   REGION R-trig
       #RTIRG_iReset(CLK := #iReset);
       #RTRIG_iFailSafe(CLK := #iFailSafe);
       #RTIRG_jog(CLK := #iJogOpen XOR #iJogClose);
       #RTIRG_auto(CLK := NOT #iMan);
       #RTRIG_iFailSafe_released(CLK := #iFailSafe);
       #RTRIG_iInterlook_released(CLK := #iInterlook);
       #RTRIG_jogOpen_released(CLK := NOT #iJogOpen);
       #RTRIG_jogClose_released(CLK := NOT #iJogClose);
   END_REGION

   REGION Timeout  

       // Quick timeout:
       // Cheak at intervals that the position moves towards the setpoint.
       // This give a quicker feedback, then the long timeout.
       IF #action <> #old.action
           OR #RTIRG_jog.Q
           OR #RTRIG_iFailSafe.Q
       THEN
           RESET_TIMER(#TONR_quckTimeoutInterval);
           #quickTimeoutLastPos := #io.in.pos;
       ELSIF #action <> #NO_ACTION AND #conf.quickTimeoutEnable THEN
           // Quick timeout in action.
           #TONR_quckTimeoutInterval.TONR(IN := #io.out.open OR #io.out.close,
                                          PT := #conf.quickTimeoutIntervalCheaks);
           IF #TONR_quckTimeoutInterval.Q THEN
               // A new interval check, now see if the valve has moved sufficient.
               #out.qucikTimeout :=
               ABS(#quickTimeoutLastPos - #io.in.pos) < #conf.qucikTimeoutMinMovement;
               RESET_TIMER(#TONR_quckTimeoutInterval);
               // Only store the old value if the valve has done progress towards the SP.
               IF #action = #OPEN AND #io.in.pos > #quickTimeoutLastPos
                   OR #action = #CLOSE AND #io.in.pos < #quickTimeoutLastPos
               THEN
                   #quickTimeoutLastPos := #io.in.pos;
               END_IF;
           END_IF;
       END_IF;

       // Long timeout:
       // Max time the valve can operate before timeout, and the valve will stop.
       #TONR_timeout.TONR(IN := #io.out.open OR #io.out.close,
                          PT := #conf.longTimeout,
                          Q => #out.longTimeout);
       // Reset timeout
       IF #RTIRG_iReset.Q
           OR #RTRIG_iFailSafe.Q
           OR #conf.autoReset AND (
           (* *)#RTIRG_jog.Q
           (* *)OR #iSP <> #old.SP AND #iMan
           (* *)OR #RTIRG_jog.Q)
       THEN
           RESET_TIMER(#TONR_timeout);
           RESET_TIMER(#TONR_quckTimeoutInterval);
           #out.qucikTimeout := false;
           #qTimeout := false;
       END_IF;
   END_REGION

   REGION Decide
       // Decide what to do ...

       // Error, timeout, failSafe and Interlook.
       IF #TONR_timeout.Q THEN
           #action := #NO_ACTION;
       ELSIF #iFailSafe THEN
           // Timeout will be reseted once if iFailSafe is activated.
           #action := #conf.feilSafeAction;
       ELSIF #iStop
           // If pos.error and there are not end-limit-switces.
           OR #io.in.posError AND (#conf.simFullyOpenWithPos OR #conf.simFullyClosedWithPos)
           OR #out.qucikTimeout
           OR #RTRIG_jogOpen_released.Q
           OR #RTRIG_jogClose_released.Q
           OR #iExternalError
       THEN
           #action := #NO_ACTION;

           // ==========================================================================
           // JOG-mode
       ELSIF #iJogOpen XOR #iJogClose THEN
           // Open or close the valve little by little. When either of the jog
           // inputs are true. This way of controlling the valve has priority
           // over setpoint (bellow).
           RESET_TIMER(#TON_regModeWait);
           IF #iJogOpen THEN
               #action := #OPEN;
           ELSIF #iJogClose THEN
               #action := #CLOSE;
           END_IF;
       ELSIF #io.in.posError THEN
           #action := #NO_ACTION;
       ELSE
           // ==========================================================================
           // SP-mode:
           // Controll the valve by a setpoint, using the feedback position to 
           // determined if the valve should open or close. SP should be given in percent.

           IF (#iSP <> #old.SP // SP has changed.
               OR #RTIRG_auto.Q // Auto has just been enabled, and the valve is out of pos.
               (* *)AND ABS(#iSP - #io.in.pos) > #conf.regModeMinOffset
               OR NOT #iMan AND ( // In auto
               (* *)#RTIRG_iReset.Q // Avoid dead lock
               (* *)OR #RTRIG_iFailSafe_released.Q
               (* *)OR #RTRIG_iInterlook_released.Q
               (* *)OR #RTRIG_jogClose_released.Q OR #RTRIG_jogOpen_released.Q )
               (* *)) AND (
               (*     *)NOT #iRegMode // Not regMode, no aditional requirements.
               (*     *)OR #TON_regModeWait.Q AND ( // A break between each move.
               (*        *)// Offset is bigger then a certain offset.
               (*        *)ABS(#iSP - #io.in.pos) > #conf.regModeMinOffset
               (*        *)// At almost closed and open, the offset requirement
               (*        *)// may not be fulfilled.
               (*        *)OR #io.in.pos > #conf.fullyOpenPosLim - #conf.endPosWithoutPreStop
               (*        *)OR #io.in.pos < #conf.endPosWithoutPreStop))
               // regMode should be used when a valve is controlled by a PID.
               // When the valve is in regMode, then there will be a time break between each 
               // movment. And there is a need a certain offset before an ajustment is done.
               // This behavior significantly prevents wear on the valve. If the valve is not
               // in regMode, then each change in SP will make the valve operate.
           THEN
               IF #iSP > #io.in.pos THEN
                   #action := #OPEN;
               ELSIF #iSP < #io.in.pos THEN
                   #action := #CLOSE;
               END_IF;
           END_IF;

           // --------------------------------------
           // SP-reached-pos:
           // 
           // In the main area where the valve operate, it will shut off the outputs, a
           // tiny bit before it reach the SP. This make the valve, stop exacly on SP.
           // In the area of almost closed and almost open this function is disable,
           // this makes sure that it's possible to open or close the valve entirly.
           #pre := SEL(G := #iSP > #conf.fullyOpenPosLim - #conf.endPosWithoutPreStop
                       OR #iSP < #conf.endPosWithoutPreStop,
                       IN0 := #conf.preStop, IN1 := 0);
           // Detect reached position
           IF #action = #OPEN AND (#io.in.pos > #iSP - #pre OR #io.in.fullyOpen)
               OR #action = #CLOSE AND (#io.in.pos < #iSP + #pre OR #io.in.fullyClosed)
           THEN
               #action := #NO_ACTION;
               RESET_TIMER(#TON_regModeWait);
           END_IF;
       END_IF;
       // In regMode this timer need to finnish before a new movement can be done.
       #TON_regModeWait.TON(IN := true,
                            PT := #conf.regModeTimeBreak);
   END_REGION

   REGION Gentle
       // If a big valve closes or open to fast, it can damage the pipes or other
       // equipment. This section make time breaks on closing or opening. 

       #gentleMode := #io.in.pos < #conf.gentleActivteLowLimit // ->
       // -> The function is only active under a ceratain position limit.
       AND (NOT #iFailSafe OR #conf.gentleAlsoOnFailSafe)
       // AlsoOnFailSafe: It's possible to disable the function for emergencies
       // by setting the value false.
       AND (#conf.gentleOpenEnable AND #action = #OPEN
       (* *)OR #conf.gentleCloseEnable AND #action = #CLOSE);    

       // The time break will increase as the valve move from the limit towards close.
       #pause := REAL_TO_DINT(#conf.gentleTimePauseBias
                              + (#io.in.pos / #conf.gentleActivteLowLimit)
                              * #conf.gentleTimePauseDelta);
       IF #gentleMode THEN
           #TON_gentle.TON(IN := true,
                           PT := SEL(G := #gentleAction, // Toggle times
                                     IN0 := #conf.gentleTimeRun,
                                     IN1 := #pause));
           IF #TON_gentle.Q THEN
               #gentleAction := NOT #gentleAction;
               RESET_TIMER(#TON_gentle); 
           END_IF;
           #action2 := SEL(G := #gentleAction, // Toggle action
                           IN0 := #action, IN1 := #NO_ACTION);
       ELSE
           RESET_TIMER(#TON_gentle);
           #gentleAction := false;
           // If the carefully-function is disabled, then just forward
           // the action value to the next stage.
           #action2 := #action;
       END_IF;
   END_REGION

   REGION Output
       // Make a smal time break when valve change direction. This make sure that
       // that both outputs are not active at the same time.
       #TP_toggleOut.TP(IN := #action2 <> #old.action2 AND #old.action2 <> #NO_ACTION,
                        PT := #conf.toggleTimeBreak);

       // Outputs
       IF #TP_toggleOut.Q THEN // A small time break.
           #io.out.open := false;
           #io.out.close := false;
       ELSIF #iFailSafe 
           OR #iJogClose OR #iJogOpen
       THEN
           // When failSafe or jog is active both the limit-switch and positon
           // signal most indicate that the valve is in correct position. This
           // in case one of the signals isn't working.
           #io.out.open := #action2 = #OPEN AND NOT #bothSensors.open;
           #io.out.close := #action2 = #CLOSE AND NOT #bothSensors.closed;
       ELSIF #iInterlook THEN
           #io.out.open := false;
           #io.out.close := false;
       ELSE
           #io.out.open := #action2 = #OPEN AND NOT #io.in.fullyOpen;
           #io.out.close := #action2 = #CLOSE AND NOT #io.in.fullyClosed;
       END_IF;
   END_REGION

   REGION Old    
       // Store values, to check if they has changed until next scan.
       #old.SP := #iSP;
       #old.action := #action;
       #old.action2 := #action2;
   END_REGION

   #qTimeout := #out.qucikTimeout OR #out.longTimeout;
END_FUNCTION_BLOCK

FUNCTION_BLOCK "motorValve"   // FB10, SCL
{ S7_Optimized_Access := 'TRUE' }
VERSION : 0.1
   VAR_INPUT
      iFeedbackPosition : Real;
      iFeddbackPosError : Bool;
      iFeedbackFullyOpen : Bool;
      iFeedbackFullyClosed : Bool;
   END_VAR
   VAR_OUTPUT
      qOpen : Bool;
      qClose : Bool := FALSE;
   END_VAR
   VAR RETAIN
      hmi : "motorValveHmiUdt";
   END_VAR
   VAR
      valve : "motorValveCtrl";
      SP : Real;
      SP_auto : Real;
   END_VAR
   VAR CONSTANT
      AUTO : SInt := 0;
      MAN_LOCAL : SInt := 1;
      MAN_REMOTE : SInt := 2;
   END_VAR
BEGIN
   // Valve with analog feedback.

   REGION Simulation
       IF #hmi.sim.enable AND NOT #valve.iFailSafe THEN
           // Simulation of input signal, not possible if in fail safe mode.
           #hmi.io.in.pos := #hmi.sim.pos;
           #hmi.io.in.posError := false;
           #hmi.io.in.fullyOpen := #hmi.sim.pos > #hmi.conf.fullyOpenPosLim;
           #hmi.io.in.fullyClosed := #hmi.sim.pos < #hmi.conf.fullyClosedPosLim;
       ELSE
           // Input mapping
           #hmi.io.in.pos := #iFeedbackPosition;
           #hmi.io.in.posError := #iFeddbackPosError;
           #hmi.io.in.fullyOpen := #iFeedbackFullyOpen;
           #hmi.io.in.fullyClosed := #iFeedbackFullyClosed;
       END_IF;
   END_REGION

   REGION Man / auto    
       IF #hmi.cmd.stop THEN
           #hmi.autoMan := #MAN_LOCAL;
       ELSIF #hmi.cmd.jogOpen XOR #hmi.cmd.jogClose THEN
           #hmi.autoMan := #MAN_LOCAL;
           #SP := #iFeedbackPosition;
       ELSIF #hmi.cmd.openFully XOR #hmi.cmd.closeFully THEN
           #hmi.autoMan := #MAN_LOCAL;
           #SP := SEL(G := #hmi.cmd.openFully, IN0 := 0, IN1 := 100);
       ELSIF #hmi.autoMan = #MAN_LOCAL THEN
           #SP := #hmi.SP;
       ELSIF #hmi.autoMan = #AUTO THEN
           #SP := #SP_auto;
           // If auto is controlled by a pid then #hmi.conf.regMode need to be enabled.
       END_IF;
       #hmi.SP := #valve.iSP := #SP_auto := #SP;
       // Forward auto or man to the valve controller.
       CASE #hmi.autoMan OF
           #MAN_LOCAL, #MAN_REMOTE:
               #valve.iMan := true;
           #AUTO:
               #valve.iMan := false;
       END_CASE;
   END_REGION

   REGION Valve controller.        
       // Main valve controller block.
       #valve(// iFailSafe
              // iInterlook
              // iRegMode
              iStop := #hmi.cmd.stop,
              iJogOpen := #hmi.cmd.jogOpen,
              iJogClose := #hmi.cmd.jogClose,
              iReset := #hmi.cmd.reset,
              qTimeout => #hmi.error.timeout,
              conf := #hmi.conf,
              io := #hmi.io);
       #qOpen := #hmi.io.out.open; // Outputs
       #qClose := #hmi.io.out.close;
   END_REGION

   REGION Position error    
       #hmi.error.posError :=
       #iFeedbackFullyOpen AND #iFeedbackFullyClosed
       OR #iFeedbackFullyOpen
       (* *)AND #iFeedbackPosition < #hmi.conf.fullyOpenPosLim - #hmi.conf.regModeMinOffset
       (* *)AND NOT #hmi.conf.simFullyOpenWithPos
       OR #iFeedbackFullyClosed
       (* *)AND #iFeedbackPosition > #hmi.conf.fullyClosedPosLim + #hmi.conf.regModeMinOffset
       (* *)AND NOT #hmi.conf.simFullyClosedWithPos;
   END_REGION

   REGION End
       // Count secounds the valve has been operating, and number of starts.
       "operatingTime"(in := #qOpen OR #qClose,
                       opr := #hmi.operatingTime);

       // Reset signals.
       #hmi.cmd.jogOpen := false;
       #hmi.cmd.jogClose := false;
       #hmi.cmd.openFully := false;
       #hmi.cmd.closeFully := false;
       #hmi.cmd.reset := false;
       #hmi.cmd.man := false;
       #hmi.cmd.auto := false;
       CASE #hmi.autoMan OF // Reset stop signal, only if in man.
           #MAN_LOCAL, #MAN_REMOTE: // If in auto, then do nothing.
               #hmi.cmd.stop := false;
       END_CASE;

       // Other signals to HMI
       #hmi.info.failSafe := #valve.iFailSafe;
       #hmi.info.interlook := #valve.iInterlook;
       #hmi.info.regMode := #valve.iRegMode;

       #hmi.sim.simByPlc := #hmi.io.simulated;
       #hmi.io.simulated := false;
   END_REGION
END_FUNCTION_BLOCK

FUNCTION_BLOCK "motorValveSimulation"   // FB20, SCL
{ S7_Optimized_Access := 'TRUE' }
VERSION : 0.1
   VAR_INPUT
      speed : Real := 1.0;
   END_VAR
   VAR_IN_OUT
      io : "motorValveIoUdt";
   END_VAR
   VAR
      old : UDInt;
      sn : UDInt;
   END_VAR
   VAR_TEMP
      t : DTL;
      "e" : Int;
   END_VAR
BEGIN
   #"e" := RD_SYS_T(#t);
   #sn := #t.NANOSECOND / 100000 + #t.SECOND * 10;

   IF #sn = #old THEN
       IF #io.out.open THEN
           #io.in.pos += #speed * 0.1;
       ELSIF #io.out.close THEN
           #io.in.pos -= #speed;
       END_IF;
   END_IF;
   #old := #sn;

   #io.in.pos := LIMIT(MN := 0, IN := #io.in.pos, MX := 100);
   #io.in.fullyOpen := #io.in.pos > 99;
   #io.in.fullyClosed := #io.in.pos < 1;

   #io.simulated := true;
END_FUNCTION_BLOCK

FUNCTION "ioGlobalMotorValveLinking" : Void   // FC24, SCL
{ S7_Optimized_Access := 'TRUE' }
VERSION : 0.1
   VAR_IN_OUT
      ioGlobal : "ioGlobal_FB";
      valve : "motorValve";
   END_VAR
BEGIN
   // Link ioGlobal with valve functions.

   // A id for each io
   #ioGlobal.z.ioIdCnt += 1;

   IF #ioGlobal.info2ioBlocks.disableAllSim THEN
       #valve.hmi.sim.enable := false;
   END_IF;
   // Count active simulations
   #ioGlobal.collectInfo.activeSimCnt +=
   BOOL_TO_UINT(#valve.hmi.sim.enable OR #valve.hmi.sim.simByPlc);

   // Count number of errors
   #ioGlobal.collectInfo.errorCnt +=
   BOOL_TO_UINT(#valve.hmi.io.in.posError OR #valve.hmi.error.timeout);
END_FUNCTION

// folder: Library/Valves/Blocks and UDT's/z Dev

FUNCTION_BLOCK "motorValveDigital"   // FB11, SCL
{ S7_Optimized_Access := 'TRUE' }
VERSION : 0.1
   VAR_INPUT
      iAction : SInt;   // 0=no-action, 1=Open, 2=Close
      iFailSafe : Bool;   // Open or close the valve entirly, set inside conf.
      iInterlook : Bool;   // Stop movement, valve will continue when input is set back false.
      iStop : Bool;   // Stop movement, also after var. is back false.
      iJogOpen : Bool;   // Move the valve towards open when true, has priority over SP.
      iJogClose : Bool;   // Move the valve towards close when true, has priority over SP.
      iReset : Bool;   // Reset timeout.
   END_VAR
   VAR_OUTPUT
      qTimeout : Bool;   // (quick and long timeout)
   END_VAR
   VAR
      action : SInt;   // 1=open, 2=close
      actionOut : SInt;
      oldAction : SInt;
      oldActionOut : SInt;
      RTIRG_iFailSafe : R_TRIG;
      RTIRG_iReset : R_TRIG;
      RTIRG_jog : R_TRIG;
      TP_toggleOut : IEC_TIMER;
      TON_gentle : IEC_TIMER;
      TONR_gentle : IEC_TIMER;
      TONR_timeout : IEC_TIMER;
      TON_regModeWait : IEC_TIMER;
      gentleAction : Bool;
   END_VAR
   VAR_TEMP
      reset : Bool;
   END_VAR
   VAR CONSTANT
      NO_ACTION : SInt := 0;
      OPEN : SInt := 1;
      CLOSE : SInt := 2;
   END_VAR
BEGIN
   // #conf - "motorValveConfUdt"
   // #io - "motorValveIoUdt"

   // Valve 

   (*

   //R-TRIG'S
   #RTIRG_iReset(CLK := #iReset);
   #RTIRG_iFailSafe(CLK := #iFailSafe); // Reset timeout once on failSafe.
   #RTIRG_jog(CLK := #iJogOpen XOR #iJogClose);

   REGION Timeout-and-reset
       // Max time the valve can operate before timeout, and the valve will stop.
       #TONR_timeout.TONR(IN := #io.out.open OR #io.out.close,
                          PT := #conf.longTimeout,
                          Q => #qTimeout);

       // Reset timeout
       IF #iJogOpen OR #iJogClose THEN
           #reset := #RTIRG_jog.Q AND (#conf.autoReset OR NOT #qTimeout);
       END_IF;
       IF #RTIRG_iReset.Q OR #RTIRG_iFailSafe.Q OR #reset THEN
           RESET_TIMER(#TONR_timeout);
           #qTimeout := false;
       END_IF;
   END_REGION

   REGION Decide
       // Error, timeout, failSafe and Interlook.
       IF #TONR_timeout.Q THEN
           #action := #NO_ACTION;
       ELSIF #iFailSafe THEN // Timeout will be reseted once if iFailSafe is activated.
           #action := #conf.feilSafeAction;
       ELSIF #iStop THEN
           #action := #NO_ACTION;
           // ==========================================================================
           // JOG-mode
       ELSIF #iJogOpen OR #iJogClose THEN
           // Open or close the valve little by little. When either of the jog
           // inputs are true. This way of controlling the valve has priority
           // over setpoint (bellow).
           RESET_TIMER(#TON_regModeWait);
           IF #iJogOpen AND #iJogClose THEN
               #action := #NO_ACTION;
           ELSIF #iJogOpen THEN
               #action := #OPEN;
           ELSIF #iJogClose THEN
               #action := #CLOSE;
           ELSE
               ;
           END_IF;
       END_IF;
   END_REGION

   REGION Gentle
       // If a big valve closes or open to fast, it can damage the pipes or other
       // equipment. This section make time breaks on closing or opening. 
       IF #io.in.pos < #conf.gentleActivteLowLimit // ->
           // -> The function is only active under a ceratain position limit.
           AND (NOT #iFailSafe OR #conf.gentleAlsoOnFailSafe)
           // AlsoOnFailSafe: It's possible to disable the function for emergencies
           // by setting the value false.
           AND (#conf.gentleOpenEnable AND #action = #OPEN
           (* *)OR #conf.gentleOpenEnable AND #action = #CLOSE)
       THEN
           #TON_gentle.PT := SEL(G := #gentleAction, // Toggle times
                                 IN0 := #conf.gentleTimeRun,
                                 IN1 := #conf.gentleTimePauseBias);
           #TON_gentle.TON(IN := true,
                           PT := #TON_gentle.PT);
           IF #TON_gentle.Q THEN
               #gentleAction := NOT #gentleAction;
               RESET_TIMER(#TON_gentle);
           END_IF;
           #actionOut := SEL(G := #gentleAction, // Toggle action
                             IN0 := #action, IN1 := #NO_ACTION);
       ELSE
           RESET_TIMER(#TON_gentle);
           #gentleAction := false;
           // If the carefully-function is disabled, then just forward
           // the action value to the next stage.
           #actionOut := #action;
       END_IF;
   END_REGION

   REGION Output
       // Make a smal time break when valve change direction. This make sure that
       // that both outputs are not active at the same time.
       #TP_toggleOut.TP(IN := #actionOut <> #oldActionOut AND #oldActionOut <> #NO_ACTION,
                        PT := #conf.toggleTimeBreak);
       // Outputs
       IF #TP_toggleOut.Q THEN
           #io.out.open := false;
           #io.out.close := false;
       ELSIF #iFailSafe THEN
           #io.out.open := #conf.feilSafeAction = #OPEN AND NOT #io.in.fullyOpen;
           #io.out.close := #conf.feilSafeAction = #CLOSE AND NOT #io.in.fullyClosed;
       ELSIF #iInterlook OR #iStop THEN
           #io.out.open := false;
           #io.out.close := false;
       ELSE
           #io.out.open := #actionOut = #OPEN AND NOT #io.in.fullyOpen;
           #io.out.close := #actionOut = #CLOSE AND NOT #io.in.fullyClosed;
       END_IF;
   END_REGION

   REGION Old
       #oldAction := #action;
       #oldActionOut := #actionOut;
   END_REGION


   // *)
END_FUNCTION_BLOCK

FUNCTION_BLOCK "motorValveAproxPos"   // FB24, SCL
{ S7_Optimized_Access := 'TRUE' }
VERSION : 0.1
   VAR_IN_OUT
      io : "motorValveIoUdt";
   END_VAR
   VAR
      conf : Struct
         maxAvoid : Real := 4.0;
      END_STRUCT;
      oldSecAndMsec10 : UInt;
      posPrT : UInt;
      "timer" : IEC_TIMER;
      first_scan : Bool := TRUE;
      RTRIG_fullyOpen : R_TRIG;
      RTRIG_fullyClosed : R_TRIG;
      rangeTime : Time;
      tries : Array[0..7] of Time;
   END_VAR
   VAR_TEMP
      "e" : Int;
      rd_sys_t : DTL;
      secAndMsec10 : UInt;
      sPos : Int;
      t : Int;
      c : Int;
      mx : Time;
      mn : Time;
   END_VAR
BEGIN
   // #io - "motorValveIoUdt"


   // For valve without position sensor. Calculate the position based on long
   // time the valve has been opening and closing.

   (* FUNCTION NOT FINISHED...

   #e := RD_SYS_T(#rd_sys_t);
   #secAndMsec10 := #rd_sys_t.SECOND * 100 + UDINT_TO_UINT(#rd_sys_t.NANOSECOND / 10000);
   #t := USINT_TO_INT( (#secAndMsec10 - #oldSecAndMsec10 + 6000) MOD 6000);
   #oldSecAndMsec10 := #secAndMsec10;

   #io.in.posError := #io.in.posError AND NOT #first_scan;

   #RTRIG_fullyOpen(CLK := #io.in.fullyOpen);
   #RTRIG_fullyClosed(CLK := #io.in.fullyClosed);

   IF #RTRIG_fullyOpen.Q OR #RTRIG_fullyClosed.Q THEN
       RESET_TIMER(#timer);
       #timer.PT := T#10m;
   END_IF;



   #c := 7 - 1;
   WHILE #c >= 0 DO
       #tries[#c + 1] := #tries[#c];
       #c -= 1;
   END_WHILE;
   #tries[0] := T#123s;

   #mn := T#24d;
   FOR #c := 1 TO 6 BY 2 DO
       #mx := MAX(IN1 := #tries[#c], IN2 := #mx);
       #mn := MIN(IN1 := #tries[#c], IN2 := #mn);
   END_FOR;
   // #mx - #mn ;

   (*IF #first_scan THEN
       #io.in.posError := true;
   END_IF;*)


   IF #io.out.open XOR #io.out.close THEN
       #sPos := SEL(G := #io.out.close, IN0 := #sPos + #t, IN1 := #sPos - #t);
   END_IF;


   // #io.in.pos

   #first_scan := false;

   *)
END_FUNCTION_BLOCK

// folder: Library/Valves/Puls valve

FUNCTION_BLOCK "pulsValve"   // FB25, SCL
{ S7_Optimized_Access := 'TRUE' }
VERSION : 0.1
   VAR_INPUT
      iOpening : Bool;
      iCloses : Bool;
      iPuls : Bool;
      iFullyOpen : Bool;
      iFullyClosed : Bool;
      iConfTimeout : Time := T#3S;
      iConfPulsesBetweenOpenAndClosed : Int;
   END_VAR
   VAR_OUTPUT
      qPos : Real;
      qUnknownPos : Bool;
   END_VAR
   VAR
      cnt : Int;
      rtrig_puls : R_TRIG;
      "timer" : IEC_TIMER;
      first_scan : Bool := TRUE;
   END_VAR
   VAR CONSTANT
      NUMBER_PULES_NOT_CONFIGERED : Int := 0;
   END_VAR
BEGIN
   // Valve position based on puls feedback 

   #rtrig_puls(CLK := #iPuls);
   #"timer".TON(IN := (#iOpening OR #iCloses) AND NOT #rtrig_puls.Q,
              PT := #iConfTimeout);
   IF #iConfPulsesBetweenOpenAndClosed = 0 // Number of pules not configured
       OR #"timer".Q
       OR #first_scan  // 
   THEN
       #qUnknownPos := true;
   ELSIF #iFullyOpen THEN
       #cnt := #iConfPulsesBetweenOpenAndClosed;
       #qUnknownPos := false;
   ELSIF #iFullyClosed THEN
       #cnt := 0;
       #qUnknownPos := false;
   ELSE
       IF #iOpening AND #iCloses THEN
           ; // No action
       ELSIF #rtrig_puls.Q THEN
           #cnt += BOOL_TO_INT(#iOpening);
           #cnt -= BOOL_TO_INT(#iCloses);
       END_IF;
   END_IF;
   #qPos := INT_TO_REAL(#cnt) / INT_TO_REAL(#iConfPulsesBetweenOpenAndClosed) * 100;
   #first_scan := false;
END_FUNCTION_BLOCK

// folder: Library/sys/Generate User Msg

FUNCTION_BLOCK "genUsrMsg"   // FB3, SCL
{ S7_Optimized_Access := 'TRUE' }
VERSION : 0.1
   VAR_INPUT
      TextID : UInt;
   END_VAR
   VAR
      TextListID : UInt;
      outgoingAlarm : Bool;   // false: Incoming alarm.
      assocValues : Array[3..10] of UInt;
      "e" : Int;
   END_VAR
   VAR_TEMP
      tmpAssocValues : AssocValues;
      c : Int;
   END_VAR
BEGIN
   // Generate user diagnostic alarms 

   // #assocValues 1 and 2 allready in use by instruction.
   FOR #c := 3 TO 10 DO
       #tmpAssocValues.Value[#c] := #assocValues[#c];
   END_FOR;

   #"e" := Gen_UsrMsg
   (Mode := 1 + BOOL_TO_UINT(#outgoingAlarm)
    ,// 1: incoming alarm. 2: outgoing alarm.
    TextID := #TextID,
   TextListID := #TextListID, // (Right click and show collom-id) 
    AssocValues := #tmpAssocValues);

   (* Assoc Values:

   "This is a usr. msg: @3I%6d@"  // Assoc val 3, 6 digits. (1st val)
   "This is an other usr. msg: @5I%6d@"  // Assoc val 5, 6 digits.

   *)
END_FUNCTION_BLOCK

FUNCTION_BLOCK "example_genUsrMsg"   // FB8, SCL
{ S7_Optimized_Access := 'TRUE' }
VERSION : 0.1
   VAR
      Gen_UsrMsg : "genUsrMsg";
      some_error : Bool;
   END_VAR
BEGIN
   #Gen_UsrMsg.TextListID := 512; // See PLC alarm text lists.

   IF #some_error THEN
       #Gen_UsrMsg(1); // Text id for this alarm 
   END_IF;
END_FUNCTION_BLOCK

// ===== library types =====

TYPE "timeFormatUdt"
   STRUCT
      OFF : SInt := 0;
      MILLISECOND : SInt := 1;
      SECOUNDS : SInt := 2;
      MINUTES : SInt := 3;
      HOURS : SInt := 4;
      DAYS : SInt := 5;
   END_STRUCT;
END_TYPE

// folder: Library/Conversion/time_to_str

FUNCTION "str::" : String   // FC30, SCL
{ S7_Optimized_Access := 'TRUE' }
VERSION : 0.1
   VAR_INPUT
      in : Time;   // Time to be converted in to string.
   END_VAR
   VAR_TEMP
      t : DTL;
      dayOrHour : Bool;
   END_VAR
BEGIN
   // Time to string.

   #t += #in; // Implicit convert to dtl.
   #t.DAY -= 1; 
   #tStr := ''; 

   IF #t.DAY <> 0 THEN
       #tStr := CONCAT(IN1 := RIGHT
                              (IN := S_CONV(#t.DAY),
                               L := 1 + BOOL_TO_INT(#t.DAY > 9)),
                              IN2 := ', ');
   END_IF;
   IF #t.HOUR <> 0 OR LEN(#tStr) <> 0 THEN
       #tStr := CONCAT(IN1 := #tStr,
                              IN2 := RIGHT
                              (IN := S_CONV(#t.HOUR),
                               L := 1 + BOOL_TO_INT(#t.HOUR > 9)),
                              IN3 := ':');
   END_IF;
   #tStr := CONCAT(IN1 := #tStr,
                          IN2 := RIGHT
                          (IN := S_CONV(#t.MINUTE),
                           L := 1 + BOOL_TO_INT(#t.MINUTE > 9)),
                          IN3 := ':');
   #tStr := CONCAT(IN1 := #tStr,
                          IN2 := RIGHT
                          (IN := S_CONV(#t.SECOND),
                           L := 1 + BOOL_TO_INT(#t.SECOND > 9)));

   // https://github.com/rexhip/
END_FUNCTION

// folder: Library/State machine

FUNCTION "sTimer" : Bool   // FC23, SCL
{ S7_Optimized_Access := 'TRUE' }
VERSION : 0.1
   VAR_INPUT
      pt : Time;
   END_VAR
   VAR_IN_OUT
      t : TON_TIME;
   END_VAR
BEGIN
   #t(IN := true, PT := #pt);
   #"timer" := #t.Q;
END_FUNCTION

// ===== library: MasterCopy "ponselMessure_ChangeMbAddr" =====

FUNCTION_BLOCK "ponselMessure_ChangeMbAddr"   // FB2, SCL
{ S7_Optimized_Access := 'TRUE' }
VERSION : 0.1
   VAR_INPUT
      current_addr : USInt;
      new_addr : UInt;
      exec : Bool := true;
   END_VAR
   VAR_OUTPUT
      Done : Bool;
      Error : Bool;
   END_VAR
   VAR_IN_OUT
      mb_query : "mb_query";
   END_VAR
   VAR_TEMP
      d : Bool;
      "e" : Bool;
   END_VAR
BEGIN
   IF #new_addr < 1 OR #new_addr > 247
       OR #new_addr = #current_addr
   THEN
       #"e" := TRUE;
   ELSIF #exec THEN
       #mb_query(mb_addr := #current_addr,
                 mode := #mb_query.c.write.holding_reg,
                 data_addr := 16#A3,
                 Done => #d,
                 Error => #"e",
                 data_ptr := #new_addr);
   END_IF;
   #Done := #d;
   #Error := #"e";
END_FUNCTION_BLOCK

// ===== library: MasterCopy "ponselMessure_changeParity" =====

FUNCTION_BLOCK "ponselMessure_changeParity"   // FB9, SCL
{ S7_Optimized_Access := 'TRUE' }
VERSION : 0.1
   VAR_INPUT
      mb_addr : USInt;
      parity : USInt;
   END_VAR
   VAR_OUTPUT
      Done : Bool;
      Error : Bool;
   END_VAR
   VAR_IN_OUT
      mb_query : "mb_query";
   END_VAR
   VAR_TEMP
      d : Bool;
      "e" : Bool;
      "word" : Word;
   END_VAR
BEGIN
   // This block isn't finnish.
   //
   IF #parity > 3 THEN
       #"e" := TRUE;
   ELSE
       CASE #parity OF
           0:  // None
               #"word".%X0 := false;
               #"word".%X1 := false;
           1:  // Odd
               #"word".%X0 := false;
               #"word".%X1 := true;
           2:  // Even
               #"word".%X0 := true;
               #"word".%X1 := false;
       END_CASE;
       (*#mb_query(mb_addr := #mb_addr,
                 mode := #mb_query.c.write.holding_reg,
                 data_addr := ,
                 Done => #d,
                 Error => #e,
                 data_ptr := #word);*)
   END_IF;
   #Done := #d;
   #Error := #"e";
END_FUNCTION_BLOCK

// ===== library: MasterCopy "ponselMessure_readSign" =====

FUNCTION_BLOCK "ponselMessure_readSign"   // FB8, SCL
{ S7_Optimized_Access := 'TRUE' }
VERSION : 0.1
   VAR_INPUT
      mb_addr : USInt;
   END_VAR
   VAR_OUTPUT
      Done : Bool;
      Error : Bool;
   END_VAR
   VAR_IN_OUT
      mb_query : "mb_query";
   END_VAR
   VAR
      signs : Array[1..3] of String[64];
   END_VAR
BEGIN
   // Read calibration signatures

   #mb_query(mb_addr := #mb_addr,
             mode := #mb_query.c.read.holding_reg,
             data_addr := 16#027e,
             data_ptr := #signs);

   IF #mb_query.Done THEN
       #Done := true;
       #Error := false;
   ELSIF #mb_query.Error THEN
       #Done := false;
       #Error := true;
   END_IF;
END_FUNCTION_BLOCK

// ===== library: MasterCopy "ponselMessure_readUnits" =====

FUNCTION_BLOCK "ponselMessure_readUnits"   // FB2, SCL
{ S7_Optimized_Access := 'TRUE' }
VERSION : 0.1
   VAR_INPUT
      mb_addr : USInt;
   END_VAR
   VAR_OUTPUT
      Done : Bool;
      Error : Bool;
   END_VAR
   VAR_IN_OUT
      mb_query : "mb_query";
   END_VAR
   VAR
      Units : Array[0..4] of String[6];
   END_VAR
BEGIN
   // 

   #mb_query(mb_addr := #mb_addr,
             mode := #mb_query.c.read.holding_reg,
             data_addr := 16#0D22,
             data_ptr := #Units);
   IF #mb_query.Done THEN
       #Done := true;
       #Error := false;
   ELSIF #mb_query.Error THEN
       #Done := false;
       #Error := true;
   END_IF;
END_FUNCTION_BLOCK

// ===== library: MasterCopy "ponselMessure_restoreDefaultCoefficients" =====

FUNCTION_BLOCK "ponselMessure_restoreDefaultCoefficients"   // FB2, SCL
{ S7_Optimized_Access := 'TRUE' }
VERSION : 0.1
   VAR_INPUT
      mb_addr : USInt;
      restorTemp : Bool;
      restorPar1 : Bool;
      restorPar2 : Bool;
      restorPar3 : Bool;
      restorPar4 : Bool;
   END_VAR
   VAR_OUTPUT
      Done : Bool;
      Error : Bool;
   END_VAR
   VAR_IN_OUT
      mb_query : "mb_query";
   END_VAR
   VAR
      "word" : Word;
      old_word : Word;
      first_scan : Bool := true;
   END_VAR
   VAR_TEMP
      d : Bool;
      "e" : Bool;
   END_VAR
BEGIN
   // Restore default calibration coefficients.

   #"word".%X0 := #restorTemp;
   #"word".%X1 := #restorPar1;
   #"word".%X2 := #restorPar2;
   #"word".%X3 := #restorPar3;
   #"word".%X4 := #restorPar4;

   IF #"word" <> #old_word AND NOT #first_scan THEN
       #mb_query(mb_addr := #mb_addr,
                 mode := #mb_query.c.write.holding_reg,
                 data_addr := 16#02,
                 Done => #d,
                 Error => #"e",
                 data_ptr := #"word");
   END_IF;
   #old_word := #"word";

   #first_scan := false;
   #Done := #d;
   #Error := #"e";
END_FUNCTION_BLOCK

// ===== library: MasterCopy "ponselMesure_calibrate" =====

FUNCTION_BLOCK "ponselMesure_calibrate"   // FB5, SCL
{ S7_Optimized_Access := 'TRUE' }
VERSION : 0.1
   VAR_INPUT
      ref_value : Real;
   END_VAR
   VAR_OUTPUT
      Done : Bool;
      Error : Bool;
   END_VAR
   VAR_IN_OUT
      mb_query : "mb_query";
      ponsel_messure : "Ponsel_mesure";
      sign : "ponselMesure_sign_udt";
   END_VAR
   VAR
      conf : Struct
         messurementsBeforeCal : USInt;
      END_STRUCT;
      mode : USInt;
      state : Int;
      oldQueryCnt : UDInt;
      error_cnt : USInt;
      dword_14c : DWord;
   END_VAR
   VAR_TEMP
      valid_value : Bool;
      tDword : DWord;
      empty : "ponselMesure_sign_udt";
   END_VAR
BEGIN
   #mb_query.mb_addr := #ponsel_messure.mb_addr;
   #mb_query.mode := #mb_query.c.write.holding_reg;
   #mb_query.Error := false;

   #Done := false;
   #Error := false;

   CASE #state OF

       10: // Wait for start signal
           #state += 1;
           #oldQueryCnt := #ponsel_messure.QueryCnt;

       11: // Do some messurements.
           #ponsel_messure.api.interval := T#2s;
           #state += BOOL_TO_INT(#ponsel_messure.QueryCnt - #oldQueryCnt >
                                 #conf.messurementsBeforeCal
                                 AND #ponsel_messure.Measurement_ok);
           #state := SEL(G := #mode = 0, IN0 := #state, IN1 := 0);
       12: // Stop messurement
           #ponsel_messure.api.wait := true;
           #state += BOOL_TO_INT(#ponsel_messure.api.idle);
       13: // Send ref. value to transmitter
           #ponsel_messure.api.wait := true; // stop messurement.
           CASE #mode OF
               1..10: // Parameters, 1 to 10
                   #mb_query.data_addr := 16#204 + (#mode - 1) * 2;
               11..12: // Temperature.
                   #mb_query.data_addr := 16#200 + (#mode - 11) * 2;
           END_CASE;
           #mb_query(data_ptr := #ref_value);
           #state += BOOL_TO_INT(#mb_query.Done);
       14: // Preperation for 14c, the word may be later written to device.
           CASE #mode OF
               1..4: // Parameter, 1 - 4  
                   #tDword.%X2 := true;
                   #tDword := SHL(IN := #tDword, N := #mode - 1);
               11: // Temperature zero and span.
                   #tDword.%X0 := true;
                   #tDword := SHL(IN := #tDword, N := #mode - 11);
           END_CASE;
           #dword_14c := #dword_14c OR #tDword; // A the bit "14c"
           #state += 1;

           // =============
           // Save

       20: // Send signature to transmitter.
           CASE #mode OF
               1..4: // Parameter, 1 - 4  // ( 16#28e - 16#27e = 16#10 )
                   #mb_query.data_addr := 16#28e + (#mode - 1) * 16#10;
               11..12: // Temperature
                   #mb_query.data_addr := 16#27e;
           END_CASE;
           #mb_query(data_ptr := #sign);
           #state += BOOL_TO_INT(#mb_query.Done);
       21: // Start use new coefficients.
           #mb_query(data_addr := 16#14c, data_ptr := #tDword);
           #state += BOOL_TO_INT(#mb_query.Done);
           // 22:
           //  #sign := #empty;
           // #state += 1;

           // =============

       30: // Chancel calibration
           #dword_14c := 0;
           #mb_query(data_addr := 16#14c, data_ptr := #dword_14c);
           #state += BOOL_TO_INT(#mb_query.Done);

           // =============

       ELSE // Reset
           #state := 0;
           #mode := 0;
           #Done := true;
           #error_cnt := 0;
   END_CASE;

   // Error handeling
   #error_cnt := BOOL_TO_USINT(#mb_query.Error);
   IF #ponsel_messure.sb.out.error
       OR #error_cnt > 3 // No more then x errors
   THEN
       #error_cnt := 0;
       #Error := true;
   END_IF;
END_FUNCTION_BLOCK

// ===== library: MasterCopy "ponselMesure_calibrateOksygen" =====

FUNCTION_BLOCK "ponselMesure_calibrateOksygen"   // FB2, SCL
{ S7_Optimized_Access := 'TRUE' }
VERSION : 0.1
   VAR_IN_OUT
      mb_query : "mb_query";
      ponsel_messure_oxygen : "Ponsel_mesure_Dissolved_oxygen";
   END_VAR
   VAR
      hmi : "ponselMesure_calibrateOxygenUdt";
      _ : Bool;
      state : Int;
      calibrate : "ponselMesure_calibrate";
   END_VAR
   VAR_TEMP
      empty : "ponselMesure_sign_udt";
   END_VAR
BEGIN
   CASE #state OF
       0:  // Wait for start signal.
           IF #hmi.startTempZeroCal THEN
               #calibrate.mode := 11; // Temperature zero (0 degrees C)
           ELSIF #hmi.startTempSpanCal THEN
               #calibrate.mode := 12; // Temperature span (25 degrees C)
           ELSIF #hmi.startOxygenZeroCal THEN
               #calibrate.mode := 1; // Oxygen zero (0 %)
           ELSIF #hmi.startOxygenSpanCal THEN
               #calibrate.mode := 4; // Oxygen span (100 %)
           ELSIF #hmi.save THEN
               #calibrate.state := 20; // Save changes.
           ELSIF #hmi.cancel THEN
               #calibrate.state := 30; // Cancel changes.
           END_IF;
           IF #calibrate.mode <> 0 THEN
               #calibrate.state := 10;
           END_IF;
           #state += 1;

       1:  // Wait for the calibration block.
           #calibrate(ref_value := #hmi.ref_value,
                      Done => #hmi.Done,
                      Error => #hmi.Error,
                      mb_query := #mb_query,
                      ponsel_messure := #ponsel_messure_oxygen.ponsel_mesure,
                      sign := #hmi.sign);
           IF #hmi.cancel THEN
               #calibrate.state := 30; // Cancel changes.
           ELSIF #calibrate.Done OR #mb_query.Error THEN
               #state := 0;
           END_IF;

   END_CASE;

   #hmi.cal_pending := #calibrate.dword_14c <> 0;

   #hmi.startTempZeroCal := false;
   #hmi.startTempSpanCal := false;
   #hmi.startOxygenZeroCal := false;
   #hmi.startOxygenSpanCal := false;
   #hmi.save := false;
   #hmi.cancel := false;
END_FUNCTION_BLOCK

// ===== library: MasterCopy "ponselMesure_calibrateOxygenUdt" =====

TYPE "ponselMesure_calibrateOxygenUdt"
   STRUCT
      startTempZeroCal : Bool;
      startTempSpanCal : Bool;
      startOxygenZeroCal : Bool;
      startOxygenSpanCal : Bool;
      save : Bool;
      cancel : Bool;
      ref_value : Real;
      sign : "ponselMesure_sign_udt";
      Done : Bool;
      Error : Bool;
      cal_pending : Bool;
   END_STRUCT;
END_TYPE

// ===== library: MasterCopy "ponselMesure_sign_udt" =====

TYPE "ponselMesure_sign_udt"
   STRUCT
      person : String[16];
      minute : String[2];
      hour : String[2];
      day : String[2];
      month : String[2];
      year : String[4];
      _ : String[4];
   END_STRUCT;
END_TYPE

(* ===== HMI "HMI_RT_2" =====
system functions are stored by id; their names below are inferred from use
connection "HMI_Connection_1": ETHERNET, S7_1200_OMS

HMI tags "Default tag table"
   "popupAnalogInTag" : WString[254] AT %DB1.DBX0.0

graphic list "@DiagnosticsStates": 0 '@Diagnostics_StateGood'; 1 '@Diagnostics_StateBad'

SlideinScreen "GraphX_Slidein_Left" 300x480
   Button "Button_4" at 43,212 size 190x34; TextOff 'Modbus'
      on Click: ActivateScreen("Modbus", 0)
   Button "Button_1" at 43,156 size 190x34; TextOff 'Home'
      on Click: ActivateScreen("Test", 0)
   Button "Button_2" at 43,268 size 190x34; TextOff 'Load balancer'
      on Click: ActivateScreen("load_balanser", 0)

SlideinScreen "GraphX_Slidein_Right" 267x480
   Button "Button_1" at 43,404 size 190x34; TextOff 'User mangement'
      on Click: ActivateScreen("UserMangement", 0)
   Button "Button_2" at 43,340 size 190x34; TextOff 'Diagnostics'
      on Click: ActivateScreen("Diagnostics", 0)
   Button "Button_3" at 43,276 size 190x34; TextOff 'Alarms'
      on Click: ActivateScreen("Alarms", 0)
   Button "Button_4" at 43,212 size 190x34; TextOff 'Test'
      on Click: ActivateScreen("Test", 0)